
       //***************************************************Setpoints Ranges***************************************************************
       IF "R-402_DB".Status.Step = 24 OR "R-402_DB".Status.Step = 25 THEN
           "Mon_R402_DB"."Min Range" := "R-402_Recipe".Temperature.SP1 - "R-402_Aux_DB"."Real"."TE-402".Temperature.MinRange;
           "Mon_R402_DB"."Max Range" := "R-402_Recipe".Temperature.SP1 + "R-402_Aux_DB"."Real"."TE-402".Temperature.MaxRange;
       ELSIF "R-402_DB".Status.Step = 26 THEN
           "Mon_R402_DB"."Min Range" := "R-402_Recipe".Temperature.SP2 - "R-402_Aux_DB"."Real"."TE-402".Temperature.MinRange;
           "Mon_R402_DB"."Max Range" := "R-402_Recipe".Temperature.SP2 + "R-402_Aux_DB"."Real"."TE-402".Temperature.MaxRange;
       ELSIF "R-402_DB".Status.Step = 27 THEN
           "Mon_R402_DB"."Min Range" := "R-402_Recipe".Temperature.SP3 - "R-402_Aux_DB"."Real"."TE-402".Temperature.MinRange;
           "Mon_R402_DB"."Max Range" := "R-402_Recipe".Temperature.SP3 + "R-402_Aux_DB"."Real"."TE-402".Temperature.MaxRange;
       END_IF;

        //***************Valves Status***************//
       "R-402_Aux_DB"."Bool".TOff := "R-402_DB".Equipments.Valves."FV-4021".TurningOff;

       //***********************************************Timers****************************************************************************//
       "R-402_Aux_DB"."Bool".HoldTimeEn := "Mon_R402_DB".ReadyToProcess AND ("R-402_SEQ_DB".S_NO = 25 OR "R-402_SEQ_DB".S_NO = 27 OR "R-402_SEQ_DB".S_NO = 29);
       "R-402_Aux_DB"."Bool".HoldTime_Reset := "R-402_DB".Status.Step = 1 OR (NOT "Mon_R402_DB".ReadyToProcess AND ("R-402_SEQ_DB".S_NO = 24 OR "R-402_SEQ_DB".S_NO = 26 OR "R-402_SEQ_DB".S_NO = 28 OR "R-402_SEQ_DB".S_NO = 30));
END_FUNCTION

FUNCTION "R-402_SEQ_FC" : Void   // FC96, LAD
{ S7_Optimized_Access := 'TRUE' }
VERSION : 0.1
   VAR_TEMP   // added for the SCL form of the ladder/FBD networks
      _w1 : Bool;
      _w2 : Bool;
      _w3 : Bool;
   END_VAR
BEGIN

REGION Network 2: Abort/Shutdown
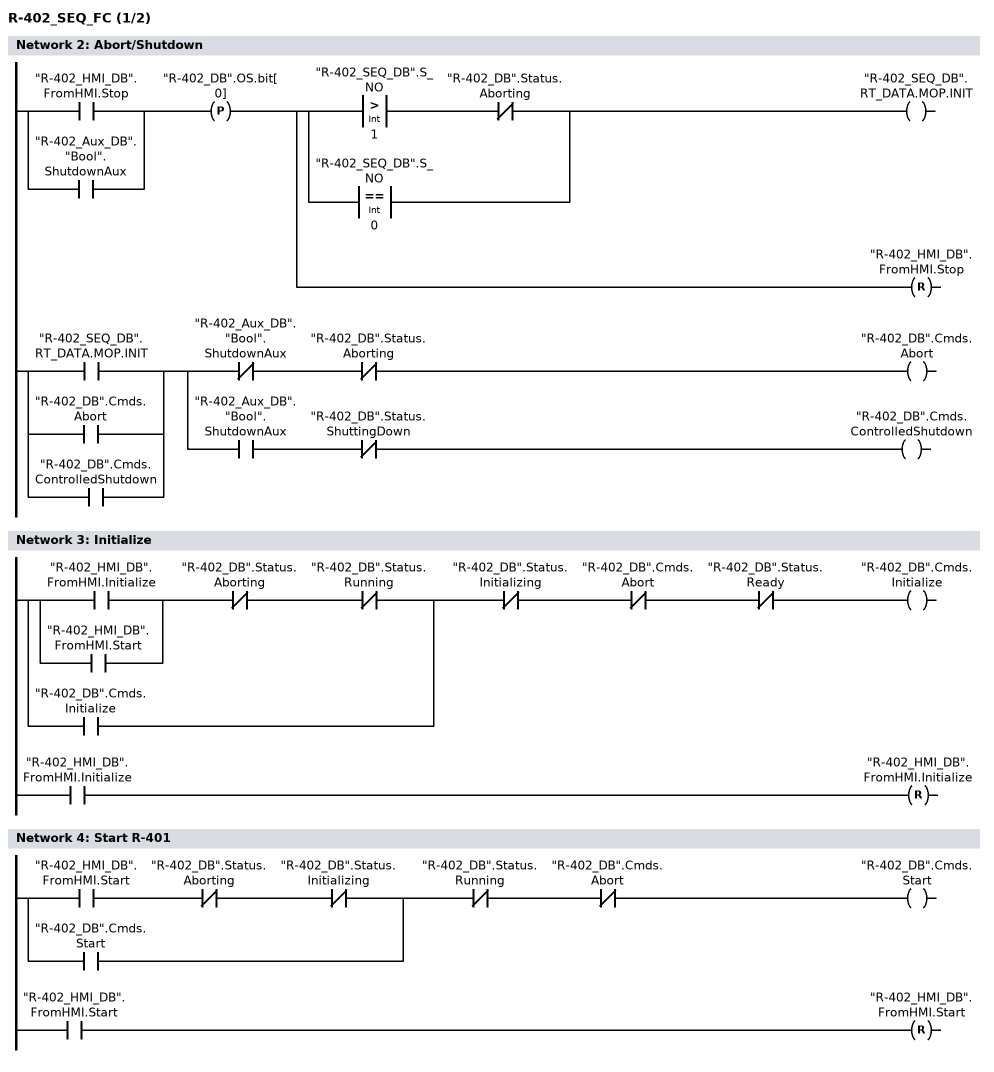
   RUNG wire#powerrail
      Contact( "R-402_HMI_DB".FromHMI.Stop )
      wire#w1
      P_Trig( "R-402_DB".OS.bit[0] )
      wire#w2
      { S7_Templates := "SrcType := Int" } GT_Contact(in1 := "R-402_SEQ_DB".S_NO, in2 := 1)
      I_Contact( "R-402_DB".Status.Aborting )
      wire#w3
      Coil( "R-402_SEQ_DB".RT_DATA.MOP.INIT )
   END_RUNG
   RUNG wire#powerrail
      Contact( "R-402_Aux_DB"."Bool".ShutdownAux )
   END_RUNG wire#w1
   RUNG wire#w2
      { S7_Templates := "SrcType := Int" } EQ_Contact(in1 := "R-402_SEQ_DB".S_NO, in2 := 0)
   END_RUNG wire#w3
   RUNG wire#w2
      R_Coil( "R-402_HMI_DB".FromHMI.Stop )
   END_RUNG
   RUNG wire#powerrail
      Contact( "R-402_SEQ_DB".RT_DATA.MOP.INIT )
      wire#w4
      I_Contact( "R-402_Aux_DB"."Bool".ShutdownAux )
      I_Contact( "R-402_DB".Status.Aborting )
      Coil( "R-402_DB".Cmds.Abort )
   END_RUNG
   RUNG wire#powerrail
      Contact( "R-402_DB".Cmds.Abort )
   END_RUNG wire#w4
   RUNG wire#powerrail
      Contact( "R-402_DB".Cmds.ControlledShutdown )
   END_RUNG wire#w4
   RUNG wire#w4
      Contact( "R-402_Aux_DB"."Bool".ShutdownAux )
      I_Contact( "R-402_DB".Status.ShuttingDown )
      Coil( "R-402_DB".Cmds.ControlledShutdown )
   END_RUNG
   // the same network as SCL:
   #_w1 := "R-402_HMI_DB".FromHMI.Stop OR "R-402_Aux_DB"."Bool".ShutdownAux;
   #_w2 := #_w1 AND NOT "R-402_DB".OS.bit[0];   // rising edge
   "R-402_DB".OS.bit[0] := #_w1;
   "R-402_SEQ_DB".RT_DATA.MOP.INIT := #_w2 AND ((("R-402_SEQ_DB".S_NO > 1) AND NOT "R-402_DB".Status.Aborting) OR ("R-402_SEQ_DB".S_NO = 0));
   IF #_w2 THEN "R-402_HMI_DB".FromHMI.Stop := FALSE; END_IF;
   #_w3 := "R-402_SEQ_DB".RT_DATA.MOP.INIT OR "R-402_DB".Cmds.Abort OR "R-402_DB".Cmds.ControlledShutdown;
   "R-402_DB".Cmds.Abort := #_w3 AND NOT "R-402_Aux_DB"."Bool".ShutdownAux AND NOT "R-402_DB".Status.Aborting;
   "R-402_DB".Cmds.ControlledShutdown := #_w3 AND "R-402_Aux_DB"."Bool".ShutdownAux AND NOT "R-402_DB".Status.ShuttingDown;
END_REGION

REGION Network 3: Initialize
   RUNG wire#powerrail
      Contact( "R-402_HMI_DB".FromHMI.Initialize )
      wire#w1
      I_Contact( "R-402_DB".Status.Aborting )
      I_Contact( "R-402_DB".Status.Running )
      wire#w2
      I_Contact( "R-402_DB".Status.Initializing )
      I_Contact( "R-402_DB".Cmds.Abort )
      I_Contact( "R-402_DB".Status.Ready )
      Coil( "R-402_DB".Cmds.Initialize )
   END_RUNG
   RUNG wire#powerrail
      Contact( "R-402_HMI_DB".FromHMI.Start )
   END_RUNG wire#w1
   RUNG wire#powerrail
      Contact( "R-402_DB".Cmds.Initialize )
   END_RUNG wire#w2
   RUNG wire#powerrail
      Contact( "R-402_HMI_DB".FromHMI.Initialize )
      R_Coil( "R-402_HMI_DB".FromHMI.Initialize )
   END_RUNG
   // the same network as SCL:
   "R-402_DB".Cmds.Initialize := ((("R-402_HMI_DB".FromHMI.Initialize OR "R-402_HMI_DB".FromHMI.Start) AND NOT "R-402_DB".Status.Aborting AND NOT "R-402_DB".Status.Running) OR "R-402_DB".Cmds.Initialize) AND NOT "R-402_DB".Status.Initializing AND NOT "R-402_DB".Cmds.Abort AND NOT "R-402_DB".Status.Ready;
   IF "R-402_HMI_DB".FromHMI.Initialize THEN "R-402_HMI_DB".FromHMI.Initialize := FALSE; END_IF;
END_REGION

REGION Network 4: Start R-401
   RUNG wire#powerrail
      Contact( "R-402_HMI_DB".FromHMI.Start )
      I_Contact( "R-402_DB".Status.Aborting )
      I_Contact( "R-402_DB".Status.Initializing )
      wire#w1
      I_Contact( "R-402_DB".Status.Running )
      I_Contact( "R-402_DB".Cmds.Abort )
      Coil( "R-402_DB".Cmds.Start )
   END_RUNG
   RUNG wire#powerrail
      Contact( "R-402_DB".Cmds.Start )
   END_RUNG wire#w1
   RUNG wire#powerrail
      Contact( "R-402_HMI_DB".FromHMI.Start )
      R_Coil( "R-402_HMI_DB".FromHMI.Start )
   END_RUNG
   // the same network as SCL:
   "R-402_DB".Cmds.Start := (("R-402_HMI_DB".FromHMI.Start AND NOT "R-402_DB".Status.Aborting AND NOT "R-402_DB".Status.Initializing) OR "R-402_DB".Cmds.Start) AND NOT "R-402_DB".Status.Running AND NOT "R-402_DB".Cmds.Abort;
   IF "R-402_HMI_DB".FromHMI.Start THEN "R-402_HMI_DB".FromHMI.Start := FALSE; END_IF;
END_REGION

REGION Network 5: Procedure Selected
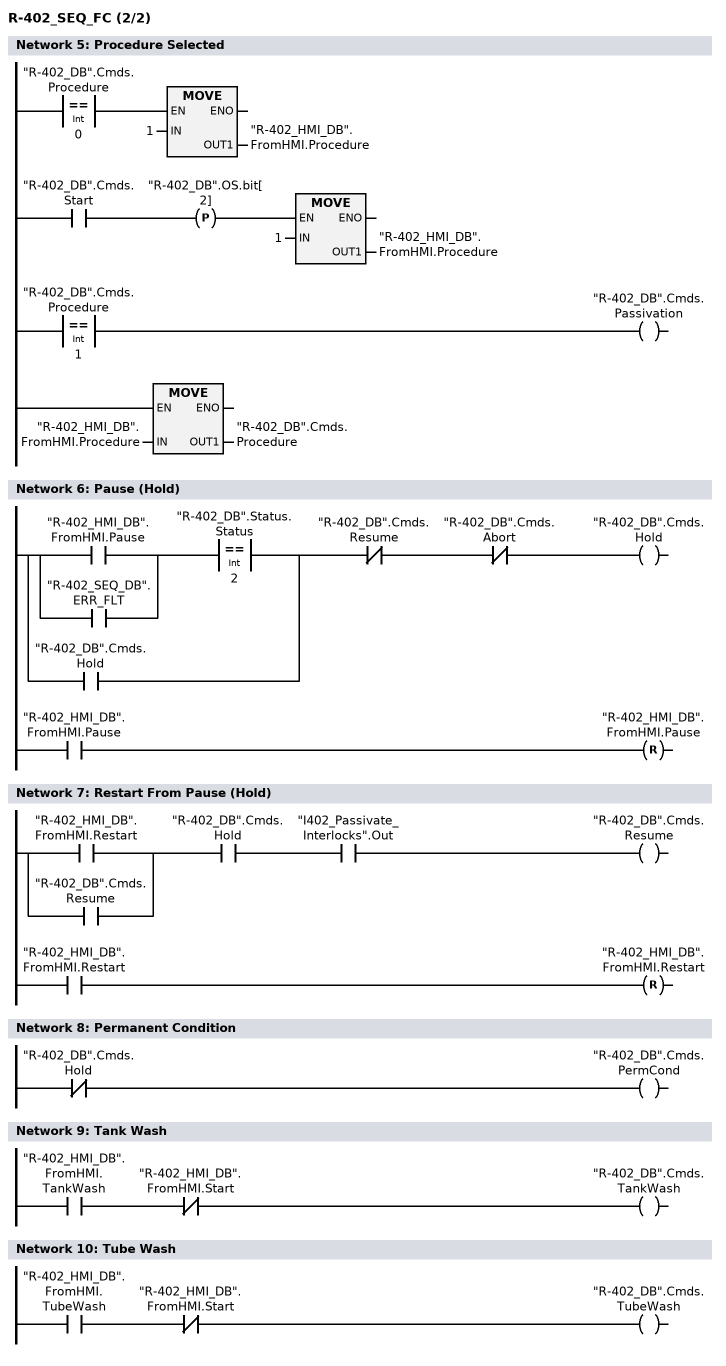
   RUNG wire#powerrail
      { S7_Templates := "SrcType := Int" } EQ_Contact(in1 := "R-402_DB".Cmds.Procedure, in2 := 0)
      Move(in := 1, out1 => "R-402_HMI_DB".FromHMI.Procedure)
   END_RUNG
   RUNG wire#powerrail
      Contact( "R-402_DB".Cmds.Start )
      P_Trig( "R-402_DB".OS.bit[2] )
      Move(in := 1, out1 => "R-402_HMI_DB".FromHMI.Procedure)
   END_RUNG
   RUNG wire#powerrail
      { S7_Templates := "SrcType := Int" } EQ_Contact(in1 := "R-402_DB".Cmds.Procedure, in2 := 1)
      Coil( "R-402_DB".Cmds.Passivation )
   END_RUNG
   RUNG wire#powerrail
      Move(in := "R-402_HMI_DB".FromHMI.Procedure, out1 => "R-402_DB".Cmds.Procedure)
   END_RUNG
   // the same network as SCL:
   IF "R-402_DB".Cmds.Procedure = 0 THEN "R-402_HMI_DB".FromHMI.Procedure := 1; END_IF;
   #_w1 := "R-402_DB".Cmds.Start AND NOT "R-402_DB".OS.bit[2];   // rising edge
   "R-402_DB".OS.bit[2] := "R-402_DB".Cmds.Start;
   IF #_w1 THEN "R-402_HMI_DB".FromHMI.Procedure := 1; END_IF;
   "R-402_DB".Cmds.Passivation := "R-402_DB".Cmds.Procedure = 1;
   "R-402_DB".Cmds.Procedure := "R-402_HMI_DB".FromHMI.Procedure;
END_REGION

REGION Network 6: Pause (Hold)
   RUNG wire#powerrail
      Contact( "R-402_HMI_DB".FromHMI.Pause )
      wire#w1
      { S7_Templates := "SrcType := Int" } EQ_Contact(in1 := "R-402_DB".Status.Status, in2 := 2)
      wire#w2
      I_Contact( "R-402_DB".Cmds.Resume )
      I_Contact( "R-402_DB".Cmds.Abort )
      Coil( "R-402_DB".Cmds.Hold )
   END_RUNG
   RUNG wire#powerrail
      Contact( "R-402_SEQ_DB".ERR_FLT )
   END_RUNG wire#w1
   RUNG wire#powerrail
      Contact( "R-402_DB".Cmds.Hold )
   END_RUNG wire#w2
   RUNG wire#powerrail
      Contact( "R-402_HMI_DB".FromHMI.Pause )
      R_Coil( "R-402_HMI_DB".FromHMI.Pause )
   END_RUNG
   // the same network as SCL:
   "R-402_DB".Cmds.Hold := ((("R-402_HMI_DB".FromHMI.Pause OR "R-402_SEQ_DB".ERR_FLT) AND ("R-402_DB".Status.Status = 2)) OR "R-402_DB".Cmds.Hold) AND NOT "R-402_DB".Cmds.Resume AND NOT "R-402_DB".Cmds.Abort;
   IF "R-402_HMI_DB".FromHMI.Pause THEN "R-402_HMI_DB".FromHMI.Pause := FALSE; END_IF;
END_REGION

REGION Network 7: Restart From Pause (Hold)
   RUNG wire#powerrail
      Contact( "R-402_HMI_DB".FromHMI.Restart )
      wire#w1
      Contact( "R-402_DB".Cmds.Hold )
      Contact( "I402_Passivate_Interlocks".Out )
      Coil( "R-402_DB".Cmds.Resume )
   END_RUNG
   RUNG wire#powerrail
      Contact( "R-402_DB".Cmds.Resume )
   END_RUNG wire#w1
   RUNG wire#powerrail
      Contact( "R-402_HMI_DB".FromHMI.Restart )
      R_Coil( "R-402_HMI_DB".FromHMI.Restart )
   END_RUNG
   // the same network as SCL:
   "R-402_DB".Cmds.Resume := ("R-402_HMI_DB".FromHMI.Restart OR "R-402_DB".Cmds.Resume) AND "R-402_DB".Cmds.Hold AND "I402_Passivate_Interlocks".Out;
   IF "R-402_HMI_DB".FromHMI.Restart THEN "R-402_HMI_DB".FromHMI.Restart := FALSE; END_IF;
END_REGION

REGION Network 8: Permanent Condition
   RUNG wire#powerrail
      I_Contact( "R-402_DB".Cmds.Hold )
      Coil( "R-402_DB".Cmds.PermCond )
   END_RUNG
   // the same network as SCL:
   "R-402_DB".Cmds.PermCond := NOT "R-402_DB".Cmds.Hold;
END_REGION

REGION Network 9: Tank Wash
   RUNG wire#powerrail
      Contact( "R-402_HMI_DB".FromHMI.TankWash )
      I_Contact( "R-402_HMI_DB".FromHMI.Start )
      Coil( "R-402_DB".Cmds.TankWash )
   END_RUNG
   // the same network as SCL:
   "R-402_DB".Cmds.TankWash := "R-402_HMI_DB".FromHMI.TankWash AND NOT "R-402_HMI_DB".FromHMI.Start;
END_REGION

REGION Network 10: Tube Wash
   RUNG wire#powerrail
      Contact( "R-402_HMI_DB".FromHMI.TubeWash )
      I_Contact( "R-402_HMI_DB".FromHMI.Start )
      Coil( "R-402_DB".Cmds.TubeWash )
   END_RUNG
   // the same network as SCL:
   "R-402_DB".Cmds.TubeWash := "R-402_HMI_DB".FromHMI.TubeWash AND NOT "R-402_HMI_DB".FromHMI.Start;
END_REGION

REGION Network 11 (SCL): Sequence Status
   IF "R-402_SEQ_DB".S_NO= 1 THEN
       "R-402_DB".Status.Status := 1; //Idle
   ELSIF ("R-402_SEQ_DB".S_NO > 1 AND "R-402_SEQ_DB".S_NO < 150) AND NOT "R-402_SEQ_DB".ERR_FLT AND NOT "R-402_DB".Cmds.Hold THEN
       "R-402_DB".Status.Status := 2; //Running
   ELSIF "R-402_SEQ_DB".S_NO >= 151 AND "R-402_SEQ_DB".S_NO <= 160 AND NOT "R-402_SEQ_DB".ERR_FLT THEN
       "R-402_DB".Status.Status := 3; // Stopping
   ELSIF  "R-402_SEQ_DB".ERR_FLT AND  ("R-402_SEQ_DB".S_NO > 1 AND "R-402_SEQ_DB".S_NO < 150) THEN
       "R-402_DB".Status.Status := 4; // Held
   ELSIF  "R-402_SEQ_DB".ERR_FLT AND  ("R-402_SEQ_DB".S_NO > 1 AND "R-402_SEQ_DB".S_NO < 150) AND "R-402_Aux_DB"."Bool".TOff  THEN
       "R-402_DB".Status.Status := 5; // Holding
   ELSE
       "R-402_DB".Status.Status := 6; // Unknown
   END_IF;

   "R-402_DB".Status.Running := ("R-402_SEQ_DB".S_NO > 3 AND "R-402_SEQ_DB".S_NO <= 150);
   "R-402_DB".Status.Initializing := ("R-402_SEQ_DB".S_NO >= 141 AND "R-402_SEQ_DB".S_NO <= 150);

   //Enable/Disable HMI Start/Stop Button
   "R-402_HMI_DB".ToHMI.EnStopButton := ("R-402_DB".Status.Status > 1) OR "R-402_DB".Status.Step = 0; //Enable HMI Stop Button
   "R-402_HMI_DB".ToHMI.EnStartButton := "R-402_DB".Status.Status = 1; //Idle
   "R-402_HMI_DB".ToHMI.EnPauseButton := "R-402_DB".Status.Status = 2; //Enable Pause Button
   "R-402_HMI_DB".ToHMI.EnRestartButton :=  "R-402_DB".Status.Status = 4; //Enable Restart Button

   //****Interlock Activated
   "R-402_HMI_DB".ToHMI.InterlockActivated := "I402_Passivate_Interlocks".Out;
END_REGION

REGION Network 12 (SCL): Sequence Step
   "R-402_DB".Status.Step := "R-402_SEQ_DB".S_NO;
END_REGION

REGION Network 13 (SCL): Sequence state (Procedure running)
   IF "R-402_SEQ_DB".S_NO = 3 OR "R-402_SEQ_DB".S_NO = 4 THEN
       "R-402_DB".Status.State := 1; //Ready
   ELSIF "R-402_SEQ_DB".S_NO >= 21 AND "R-402_SEQ_DB".S_NO <= 60 THEN
       "R-402_DB".Status.State := 2; //Mixing 
   ELSIF "R-402_SEQ_DB".S_NO >= 61 AND "R-402_SEQ_DB".S_NO <= 80 THEN
       "R-402_DB".Status.State := 3; //Pouring
   ELSIF "R-402_SEQ_DB".S_NO >= 141 AND "R-402_SEQ_DB".S_NO <= 150 THEN
       "R-402_DB".Status.State := 4; //Initializing
   ELSIF "R-402_SEQ_DB".S_NO >= 151 AND "R-402_SEQ_DB".S_NO <= 160 THEN
       "R-402_DB".Status.State := 5; //Aborting
   ELSE
       "R-402_DB".Status.State := 0;
   END_IF;
END_REGION

REGION Network 14: Sequence State
END_REGION
END_FUNCTION

// folder: Timers

FUNCTION "TIMER_FC" : Void   // FC19, LAD
{ S7_Optimized_Access := 'TRUE' }
VERSION : 0.1
   VAR_TEMP
      Reactor1ToCentrifuge : Bool;
      Reactor2ToCentrifuge : Bool;
   END_VAR
BEGIN

REGION Network 1: New Logic Timers T-101
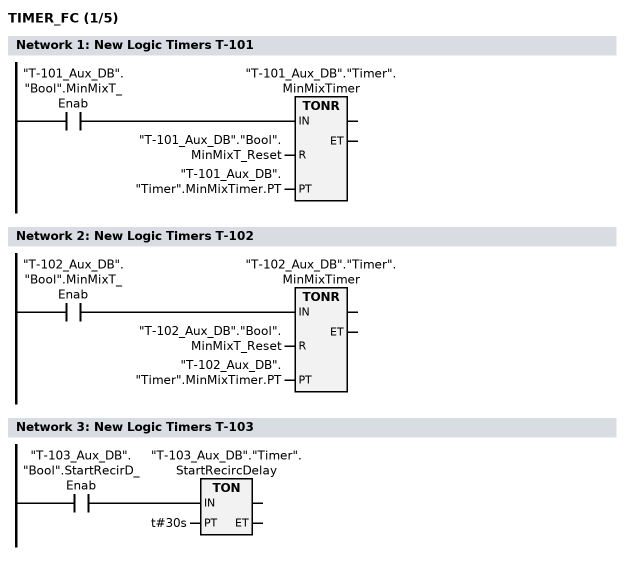
   "T-101_Aux_DB"."Timer".MinMixTimer.TONR(IN := "T-101_Aux_DB"."Bool".MinMixT_Enab,
                           R := "T-101_Aux_DB"."Bool".MinMixT_Reset,
                           PT := "T-101_Aux_DB"."Timer".MinMixTimer.PT);
END_REGION

REGION Network 2: New Logic Timers T-102
   "T-102_Aux_DB"."Timer".MinMixTimer.TONR(IN := "T-102_Aux_DB"."Bool".MinMixT_Enab,
                           R := "T-102_Aux_DB"."Bool".MinMixT_Reset,
                           PT := "T-102_Aux_DB"."Timer".MinMixTimer.PT);
END_REGION

REGION Network 3: New Logic Timers T-103
   "T-103_Aux_DB"."Timer".StartRecircDelay.TON(IN := "T-103_Aux_DB"."Bool".StartRecirD_Enab, PT := t#30s);
END_REGION

REGION Network 4: New Logic Timers R-201
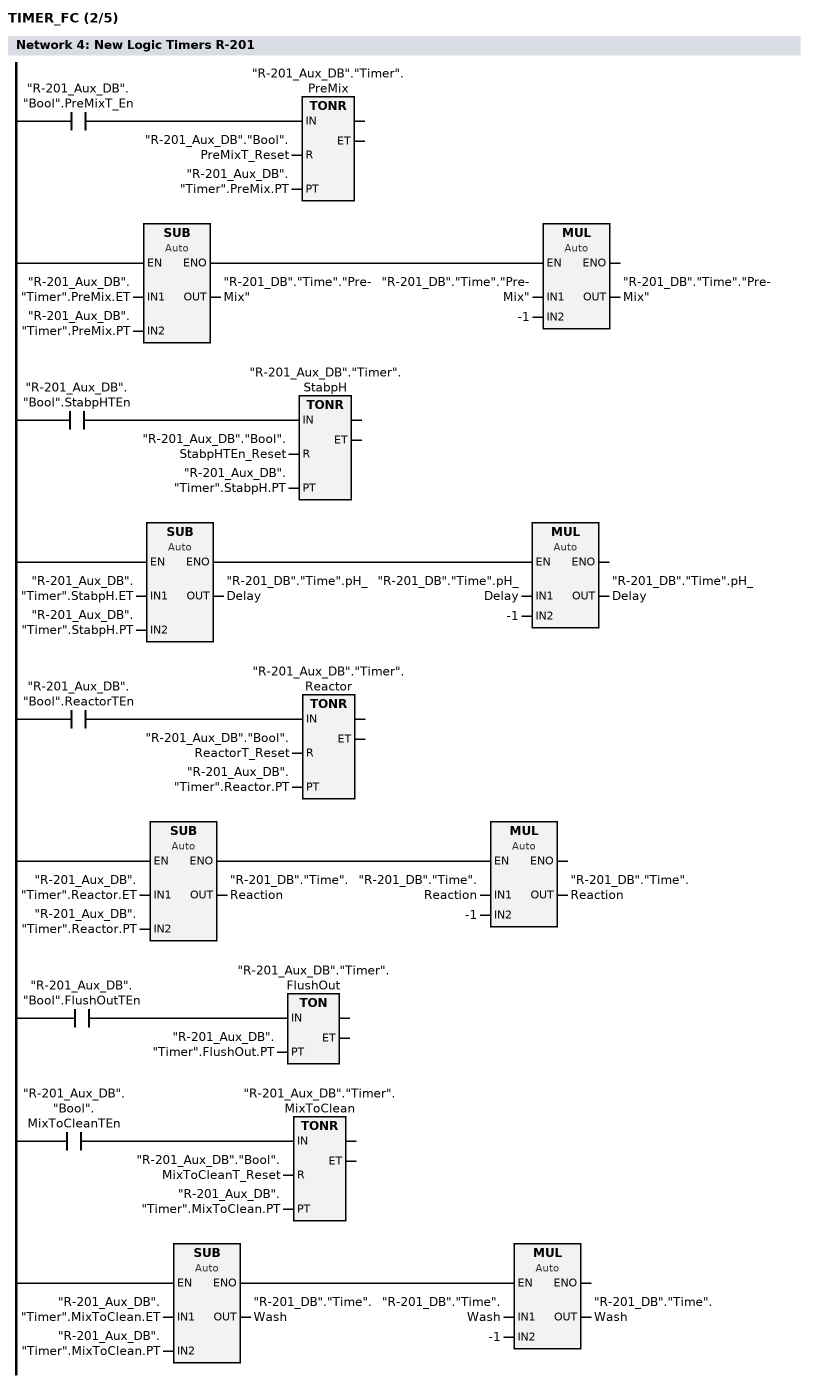
   // ENO of a box is taken as its EN; it also drops when the box reports an error
   "R-201_Aux_DB"."Timer".PreMix.TONR(IN := "R-201_Aux_DB"."Bool".PreMixT_En,
                           R := "R-201_Aux_DB"."Bool".PreMixT_Reset,
                           PT := "R-201_Aux_DB"."Timer".PreMix.PT);
   "R-201_DB"."Time"."Pre-Mix" := "R-201_Aux_DB"."Timer".PreMix.ET - "R-201_Aux_DB"."Timer".PreMix.PT;
   "R-201_DB"."Time"."Pre-Mix" := "R-201_DB"."Time"."Pre-Mix" * (-1);
   "R-201_Aux_DB"."Timer".StabpH.TONR(IN := "R-201_Aux_DB"."Bool".StabpHTEn,
                           R := "R-201_Aux_DB"."Bool".StabpHTEn_Reset,
                           PT := "R-201_Aux_DB"."Timer".StabpH.PT);
   "R-201_DB"."Time".pH_Delay := "R-201_Aux_DB"."Timer".StabpH.ET - "R-201_Aux_DB"."Timer".StabpH.PT;
   "R-201_DB"."Time".pH_Delay := "R-201_DB"."Time".pH_Delay * (-1);
   "R-201_Aux_DB"."Timer".Reactor.TONR(IN := "R-201_Aux_DB"."Bool".ReactorTEn,
                           R := "R-201_Aux_DB"."Bool".ReactorT_Reset,
                           PT := "R-201_Aux_DB"."Timer".Reactor.PT);
   "R-201_DB"."Time".Reaction := "R-201_Aux_DB"."Timer".Reactor.ET - "R-201_Aux_DB"."Timer".Reactor.PT;
   "R-201_DB"."Time".Reaction := "R-201_DB"."Time".Reaction * (-1);
   "R-201_Aux_DB"."Timer".FlushOut.TON(IN := "R-201_Aux_DB"."Bool".FlushOutTEn,
                           PT := "R-201_Aux_DB"."Timer".FlushOut.PT);
   "R-201_Aux_DB"."Timer".MixToClean.TONR(IN := "R-201_Aux_DB"."Bool".MixToCleanTEn,
                           R := "R-201_Aux_DB"."Bool".MixToCleanT_Reset,
                           PT := "R-201_Aux_DB"."Timer".MixToClean.PT);
   "R-201_DB"."Time".Wash := "R-201_Aux_DB"."Timer".MixToClean.ET - "R-201_Aux_DB"."Timer".MixToClean.PT;
   "R-201_DB"."Time".Wash := "R-201_DB"."Time".Wash * (-1);
END_REGION

REGION Network 5: New Logic Timers R-202
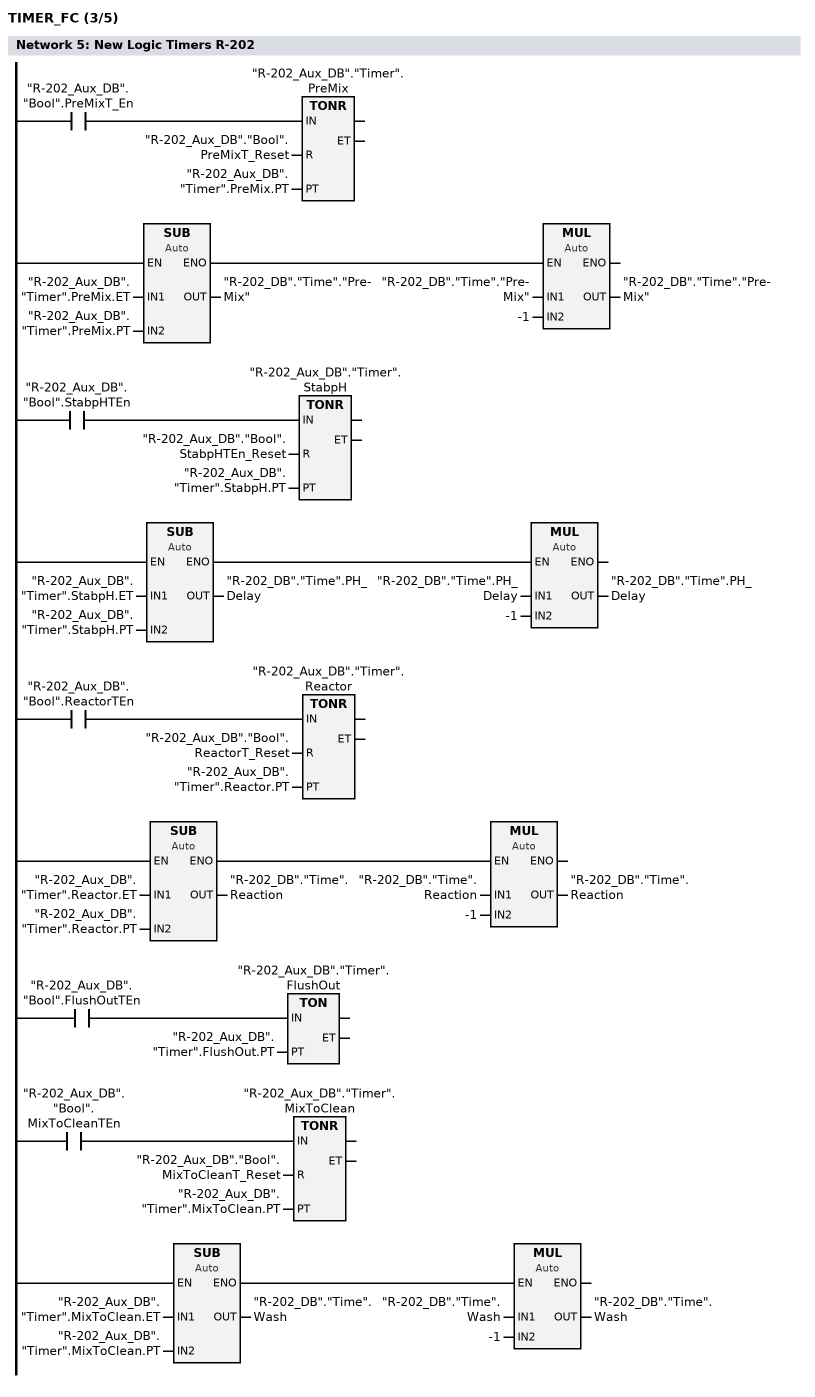
   // ENO of a box is taken as its EN; it also drops when the box reports an error
   "R-202_Aux_DB"."Timer".PreMix.TONR(IN := "R-202_Aux_DB"."Bool".PreMixT_En,
                           R := "R-202_Aux_DB"."Bool".PreMixT_Reset,
                           PT := "R-202_Aux_DB"."Timer".PreMix.PT);
   "R-202_DB"."Time"."Pre-Mix" := "R-202_Aux_DB"."Timer".PreMix.ET - "R-202_Aux_DB"."Timer".PreMix.PT;
   "R-202_DB"."Time"."Pre-Mix" := "R-202_DB"."Time"."Pre-Mix" * (-1);
   "R-202_Aux_DB"."Timer".StabpH.TONR(IN := "R-202_Aux_DB"."Bool".StabpHTEn,
                           R := "R-202_Aux_DB"."Bool".StabpHTEn_Reset,
                           PT := "R-202_Aux_DB"."Timer".StabpH.PT);
   "R-202_DB"."Time".PH_Delay := "R-202_Aux_DB"."Timer".StabpH.ET - "R-202_Aux_DB"."Timer".StabpH.PT;
   "R-202_DB"."Time".PH_Delay := "R-202_DB"."Time".PH_Delay * (-1);
   "R-202_Aux_DB"."Timer".Reactor.TONR(IN := "R-202_Aux_DB"."Bool".ReactorTEn,
                           R := "R-202_Aux_DB"."Bool".ReactorT_Reset,
                           PT := "R-202_Aux_DB"."Timer".Reactor.PT);
   "R-202_DB"."Time".Reaction := "R-202_Aux_DB"."Timer".Reactor.ET - "R-202_Aux_DB"."Timer".Reactor.PT;
   "R-202_DB"."Time".Reaction := "R-202_DB"."Time".Reaction * (-1);
   "R-202_Aux_DB"."Timer".FlushOut.TON(IN := "R-202_Aux_DB"."Bool".FlushOutTEn,
                           PT := "R-202_Aux_DB"."Timer".FlushOut.PT);
   "R-202_Aux_DB"."Timer".MixToClean.TONR(IN := "R-202_Aux_DB"."Bool".MixToCleanTEn,
                           R := "R-202_Aux_DB"."Bool".MixToCleanT_Reset,
                           PT := "R-202_Aux_DB"."Timer".MixToClean.PT);
   "R-202_DB"."Time".Wash := "R-202_Aux_DB"."Timer".MixToClean.ET - "R-202_Aux_DB"."Timer".MixToClean.PT;
   "R-202_DB"."Time".Wash := "R-202_DB"."Time".Wash * (-1);
END_REGION

REGION Network 6: New Logic Timers Centrifuge
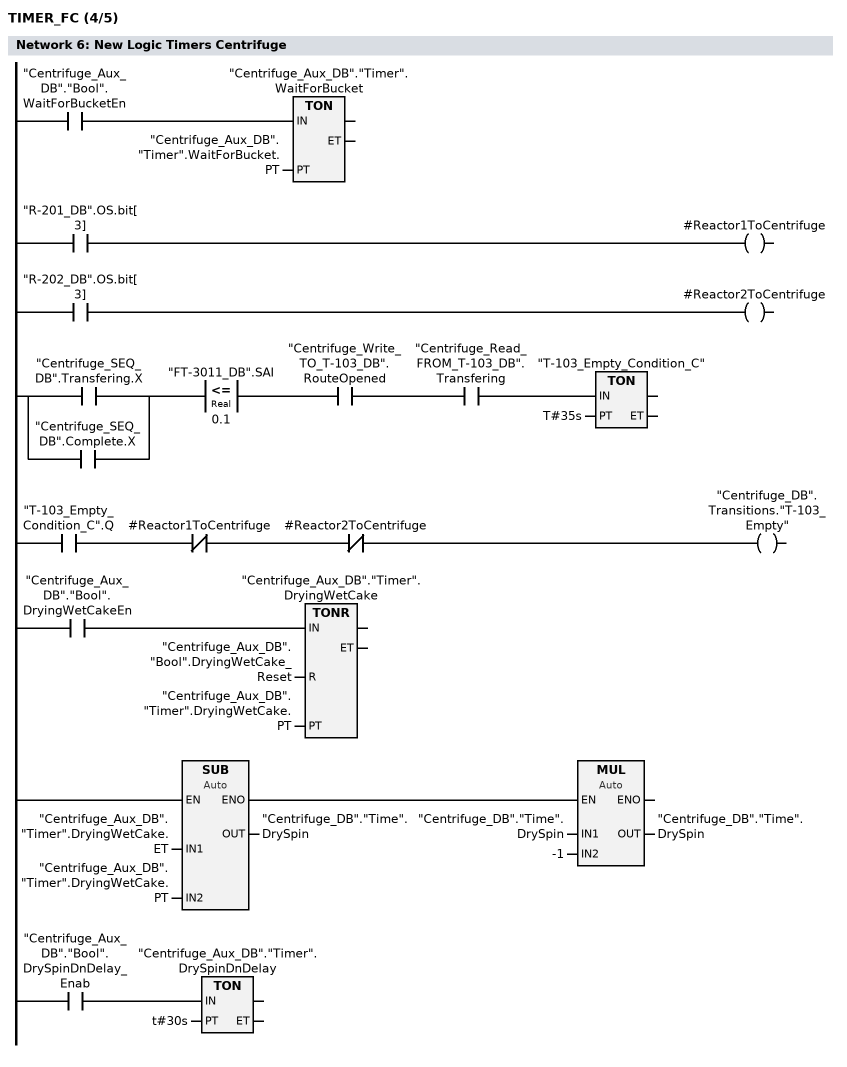
   // ENO of a box is taken as its EN; it also drops when the box reports an error
   "Centrifuge_Aux_DB"."Timer".WaitForBucket.TON(IN := "Centrifuge_Aux_DB"."Bool".WaitForBucketEn,
                           PT := "Centrifuge_Aux_DB"."Timer".WaitForBucket.PT);
   #Reactor1ToCentrifuge := "R-201_DB".OS.bit[3];
   #Reactor2ToCentrifuge := "R-202_DB".OS.bit[3];
   "T-103_Empty_Condition_C".TON(IN := ("Centrifuge_SEQ_DB".Transfering.X OR "Centrifuge_SEQ_DB".Complete.X) AND ("FT-3011_DB".SAI <= 0.1) AND "Centrifuge_Write_TO_T-103_DB".RouteOpened AND "Centrifuge_Read_FROM_T-103_DB".Transfering,
                           PT := T#35s);
   "Centrifuge_DB".Transitions."T-103_Empty" := "T-103_Empty_Condition_C".Q AND NOT #Reactor1ToCentrifuge AND NOT #Reactor2ToCentrifuge;
   "Centrifuge_Aux_DB"."Timer".DryingWetCake.TONR(IN := "Centrifuge_Aux_DB"."Bool".DryingWetCakeEn,
                           R := "Centrifuge_Aux_DB"."Bool".DryingWetCake_Reset,
                           PT := "Centrifuge_Aux_DB"."Timer".DryingWetCake.PT);
   "Centrifuge_DB"."Time".DrySpin := "Centrifuge_Aux_DB"."Timer".DryingWetCake.ET - "Centrifuge_Aux_DB"."Timer".DryingWetCake.PT;
   "Centrifuge_DB"."Time".DrySpin := "Centrifuge_DB"."Time".DrySpin * (-1);
   "Centrifuge_Aux_DB"."Timer".DrySpinDnDelay.TON(IN := "Centrifuge_Aux_DB"."Bool".DrySpinDnDelay_Enab,
                           PT := t#30s);
END_REGION

REGION Network 7: Calcination Timers
   // """Was Located in the reset of the Calcination timer"""
   // "Calcination_GRAPH_DB"."R-401 Calcination".RESET
   // ***This value was located in the PT TONR***
   // "Calcination_GRAPH_DB"."R-401 Calcination".TIMER.Calcination.PT
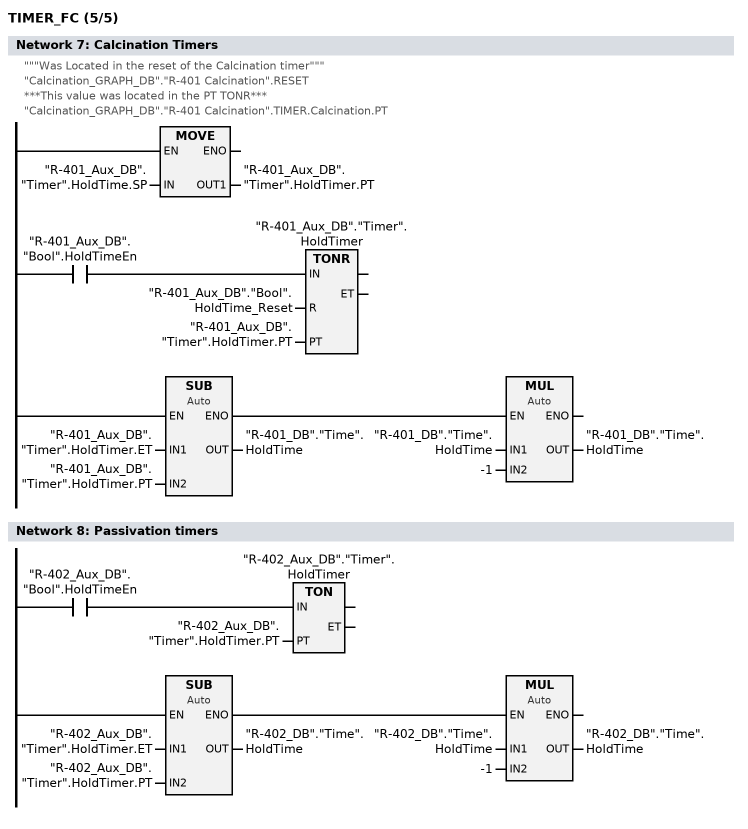
   // ENO of a box is taken as its EN; it also drops when the box reports an error
   "R-401_Aux_DB"."Timer".HoldTimer.PT := "R-401_Aux_DB"."Timer".HoldTime.SP;
   "R-401_Aux_DB"."Timer".HoldTimer.TONR(IN := "R-401_Aux_DB"."Bool".HoldTimeEn,
                           R := "R-401_Aux_DB"."Bool".HoldTime_Reset,
                           PT := "R-401_Aux_DB"."Timer".HoldTimer.PT);
   "R-401_DB"."Time".HoldTime := "R-401_Aux_DB"."Timer".HoldTimer.ET - "R-401_Aux_DB"."Timer".HoldTimer.PT;
   "R-401_DB"."Time".HoldTime := "R-401_DB"."Time".HoldTime * (-1);
END_REGION

REGION Network 8: Passivation timers
   // ENO of a box is taken as its EN; it also drops when the box reports an error
   "R-402_Aux_DB"."Timer".HoldTimer.TON(IN := "R-402_Aux_DB"."Bool".HoldTimeEn,
                           PT := "R-402_Aux_DB"."Timer".HoldTimer.PT);
   "R-402_DB"."Time".HoldTime := "R-402_Aux_DB"."Timer".HoldTimer.ET - "R-402_Aux_DB"."Timer".HoldTimer.PT;
   "R-402_DB"."Time".HoldTime := "R-402_DB"."Time".HoldTime * (-1);
END_REGION
END_FUNCTION

// folder: Timers/Totalizer

FUNCTION "Totalizers" : Void   // FC10, LAD
{ S7_Optimized_Access := 'TRUE' }
VERSION : 0.1
   VAR_TEMP   // added for the SCL form of the ladder/FBD networks
      _w1 : Bool;
      _w2 : Bool;
      _w3 : Bool;
      _w4 : Bool;
   END_VAR
BEGIN

REGION Network 1: FT-1041: T-101Water Flow Totalizer
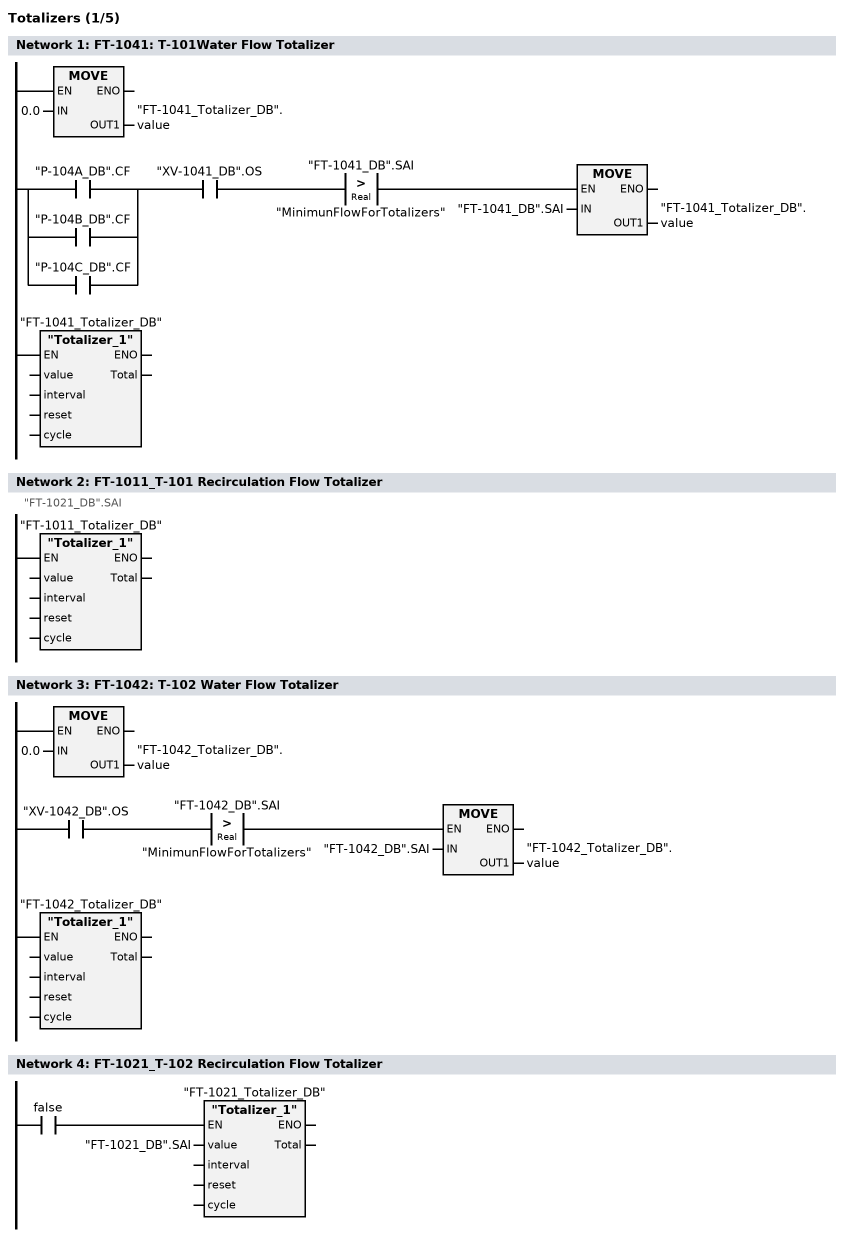
   RUNG wire#powerrail
      { S7_GenerateENO := "TRUE" } Move(in := 0.0, out1 => "FT-1041_Totalizer_DB".value)
   END_RUNG
   RUNG wire#powerrail
      Contact( "P-104A_DB".CF )
      wire#w1
      Contact( "XV-1041_DB".OS )
      { S7_Templates := "SrcType := Real" } GT_Contact(in1 := "FT-1041_DB".SAI, in2 := "MinimunFlowForTotalizers")
      { S7_GenerateENO := "TRUE" } Move(in := "FT-1041_DB".SAI, out1 => "FT-1041_Totalizer_DB".value)
   END_RUNG
   RUNG wire#powerrail
      Contact( "P-104B_DB".CF )
   END_RUNG wire#w1
   RUNG wire#powerrail
      Contact( "P-104C_DB".CF )
   END_RUNG wire#w1
   RUNG wire#powerrail
      "FT-1041_Totalizer_DB"(value :=, interval :=, reset :=, cycle :=, Total =>)
   END_RUNG
   // the same network as SCL:
   "FT-1041_Totalizer_DB".value := 0.0;
   IF ("P-104A_DB".CF OR "P-104B_DB".CF OR "P-104C_DB".CF) AND "XV-1041_DB".OS AND ("FT-1041_DB".SAI > "MinimunFlowForTotalizers") THEN
       "FT-1041_Totalizer_DB".value := "FT-1041_DB".SAI;
   END_IF;
   "FT-1041_Totalizer_DB"();   // "Totalizer_1"
END_REGION

REGION Network 2: FT-1011_T-101 Recirculation Flow Totalizer
   // "FT-1021_DB".SAI
   RUNG wire#powerrail
      "FT-1011_Totalizer_DB"(value :=, interval :=, reset :=, cycle :=, Total =>)
   END_RUNG
   // the same network as SCL:
   "FT-1011_Totalizer_DB"();   // "Totalizer_1"
END_REGION

REGION Network 3: FT-1042: T-102 Water Flow Totalizer
   RUNG wire#powerrail
      { S7_GenerateENO := "TRUE" } Move(in := 0.0, out1 => "FT-1042_Totalizer_DB".value)
   END_RUNG
   RUNG wire#powerrail
      Contact( "XV-1042_DB".OS )
      { S7_Templates := "SrcType := Real" } GT_Contact(in1 := "FT-1042_DB".SAI, in2 := "MinimunFlowForTotalizers")
      { S7_GenerateENO := "TRUE" } Move(in := "FT-1042_DB".SAI, out1 => "FT-1042_Totalizer_DB".value)
   END_RUNG
   RUNG wire#powerrail
      "FT-1042_Totalizer_DB"(value :=, interval :=, reset :=, cycle :=, Total =>)
   END_RUNG
   // the same network as SCL:
   "FT-1042_Totalizer_DB".value := 0.0;
   IF "XV-1042_DB".OS AND ("FT-1042_DB".SAI > "MinimunFlowForTotalizers") THEN
       "FT-1042_Totalizer_DB".value := "FT-1042_DB".SAI;
   END_IF;
   "FT-1042_Totalizer_DB"();   // "Totalizer_1"
END_REGION

REGION Network 4: FT-1021_T-102 Recirculation Flow Totalizer
   RUNG wire#powerrail
      Contact( false )
      "FT-1021_Totalizer_DB"(value := "FT-1021_DB".SAI, interval :=, reset :=, cycle :=, Total =>)
   END_RUNG
   // the same network as SCL:
   IF false THEN
       "FT-1021_Totalizer_DB"(value := "FT-1021_DB".SAI);   // "Totalizer_1"
   END_IF;
END_REGION

REGION Network 5: FT-1043:R-201 Water Flow Totalizer
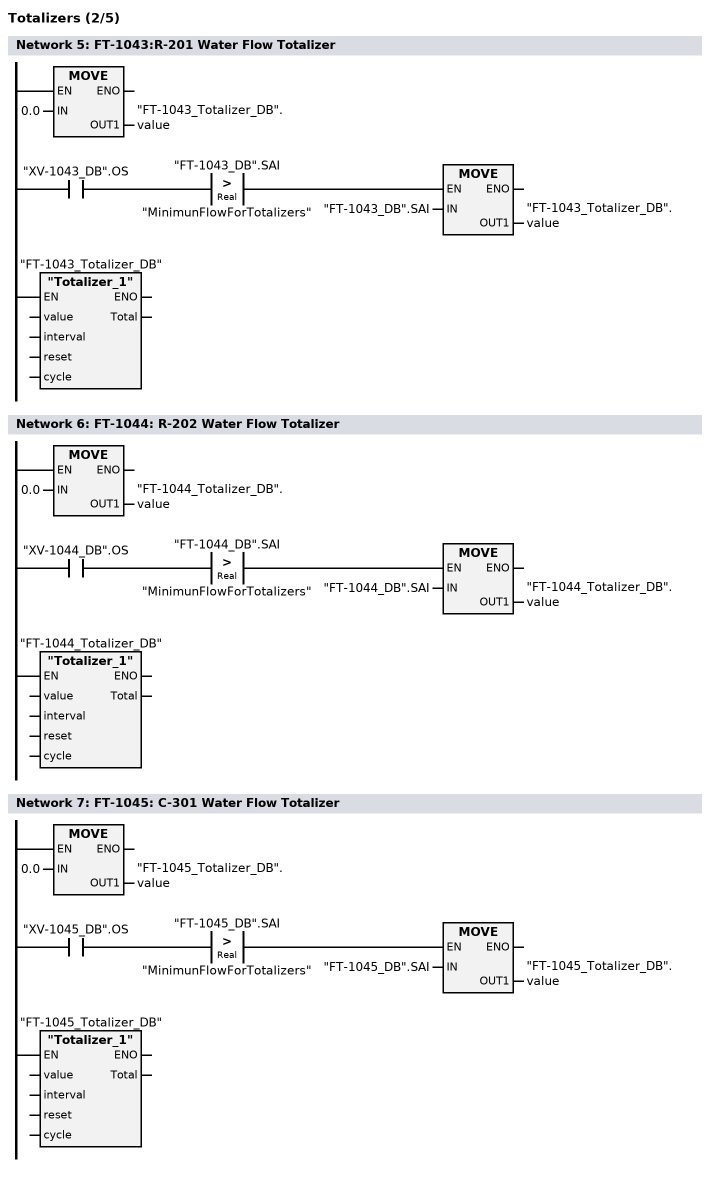
   RUNG wire#powerrail
      { S7_GenerateENO := "TRUE" } Move(in := 0.0, out1 => "FT-1043_Totalizer_DB".value)
   END_RUNG
   RUNG wire#powerrail
      Contact( "XV-1043_DB".OS )
      { S7_Templates := "SrcType := Real" } GT_Contact(in1 := "FT-1043_DB".SAI, in2 := "MinimunFlowForTotalizers")
      { S7_GenerateENO := "TRUE" } Move(in := "FT-1043_DB".SAI, out1 => "FT-1043_Totalizer_DB".value)
   END_RUNG
   RUNG wire#powerrail
      "FT-1043_Totalizer_DB"(value :=, interval :=, reset :=, cycle :=, Total =>)
   END_RUNG
   // the same network as SCL:
   "FT-1043_Totalizer_DB".value := 0.0;
   IF "XV-1043_DB".OS AND ("FT-1043_DB".SAI > "MinimunFlowForTotalizers") THEN
       "FT-1043_Totalizer_DB".value := "FT-1043_DB".SAI;
   END_IF;
   "FT-1043_Totalizer_DB"();   // "Totalizer_1"
END_REGION

REGION Network 6: FT-1044: R-202 Water Flow Totalizer
   RUNG wire#powerrail
      { S7_GenerateENO := "TRUE" } Move(in := 0.0, out1 => "FT-1044_Totalizer_DB".value)
   END_RUNG
   RUNG wire#powerrail
      Contact( "XV-1044_DB".OS )
      { S7_Templates := "SrcType := Real" } GT_Contact(in1 := "FT-1044_DB".SAI, in2 := "MinimunFlowForTotalizers")
      { S7_GenerateENO := "TRUE" } Move(in := "FT-1044_DB".SAI, out1 => "FT-1044_Totalizer_DB".value)
   END_RUNG
   RUNG wire#powerrail
      "FT-1044_Totalizer_DB"(value :=, interval :=, reset :=, cycle :=, Total =>)
   END_RUNG
   // the same network as SCL:
   "FT-1044_Totalizer_DB".value := 0.0;
   IF "XV-1044_DB".OS AND ("FT-1044_DB".SAI > "MinimunFlowForTotalizers") THEN
       "FT-1044_Totalizer_DB".value := "FT-1044_DB".SAI;
   END_IF;
   "FT-1044_Totalizer_DB"();   // "Totalizer_1"
END_REGION

REGION Network 7: FT-1045: C-301 Water Flow Totalizer
   RUNG wire#powerrail
      { S7_GenerateENO := "TRUE" } Move(in := 0.0, out1 => "FT-1045_Totalizer_DB".value)
   END_RUNG
   RUNG wire#powerrail
      Contact( "XV-1045_DB".OS )
      { S7_Templates := "SrcType := Real" } GT_Contact(in1 := "FT-1045_DB".SAI, in2 := "MinimunFlowForTotalizers")
      { S7_GenerateENO := "TRUE" } Move(in := "FT-1045_DB".SAI, out1 => "FT-1045_Totalizer_DB".value)
   END_RUNG
   RUNG wire#powerrail
      "FT-1045_Totalizer_DB"(value :=, interval :=, reset :=, cycle :=, Total =>)
   END_RUNG
   // the same network as SCL:
   "FT-1045_Totalizer_DB".value := 0.0;
   IF "XV-1045_DB".OS AND ("FT-1045_DB".SAI > "MinimunFlowForTotalizers") THEN
       "FT-1045_Totalizer_DB".value := "FT-1045_DB".SAI;
   END_IF;
   "FT-1045_Totalizer_DB"();   // "Totalizer_1"
END_REGION

